// TIA Portal project "Respirator2020_V16" (V16) (continued)
REGION Network 6: Volume/Minute Alarms / Minute Volume Alarms
   RUNG wire#powerrail
      "DirectAnalog_DB_VolumeMinute"(Pulse := "Clock_1Hz", ACK := "Operation".GeneralAck, Reset := "Operation".GeneralReset, Interlock := "Operation".InterlockVolMinute, Delay := T#1000ms, Factor := "OperatingParameters".VolumeMinFactor, AnalogInput := "DataValues".VolumeMinuteValue, SetpointPreAlarmHI := "ProcessData".VolumeMinSetpointPreAlarmHI, SetpointAlarmHI := "ProcessData".VolumeMinSetpointAlarmHI, SetpointPreAlarmLOW := "ProcessData".VolumeMinSetpointPreAlarmLOW, SetpointAlarmLOW := "ProcessData".VolumeMinSetpointAlarmLOW, HysteresisHI := "ProcessData".VolumeMinHysteresisHI, HysteresisLOW := "ProcessData".VolumeMinHysteresisLOW, DisplayPreAlarmHI => "AlarmsRaw".VolumeMinuteDisplayPreAlarmHI, InterlockPreAlarmHI => "AlarmsRaw".VolumeMinuteInterlockPreAlarmHI, DisplayAlarmHI => "AlarmsRaw".VolumeMinuteDisplayAlarmHI, InterlockAlarmHI => "AlarmsRaw".VolumeMinuteInterlockAlarmHI, DisplayPreAlarmLOW => "AlarmsRaw".VolumeMinuteDisplayPreAlarmLOW, InterlockPreAlarmLOW => "AlarmsRaw".VolumeMinuteInterlockPreAlarmLOW, DisplayAlarmLOW => "AlarmsRaw".VolumeMinuteDisplayAlarmLOW, InterlockAlarmLOW => "AlarmsRaw".VolumeMinuteInterlockAlarmLOW, CovertedOutput =>, CalcHysterisHI =>, CalcHysteresisLOW =>, DATOS =>)
   END_RUNG
   // the same network as SCL:
   "DirectAnalog_DB_VolumeMinute"(Pulse := "Clock_1Hz",   // "DirectAnalog"
                           ACK := "Operation".GeneralAck,
                           Reset := "Operation".GeneralReset,
                           Interlock := "Operation".InterlockVolMinute,
                           Delay := T#1000ms,
                           Factor := "OperatingParameters".VolumeMinFactor,
                           AnalogInput := "DataValues".VolumeMinuteValue,
                           SetpointPreAlarmHI := "ProcessData".VolumeMinSetpointPreAlarmHI,
                           SetpointAlarmHI := "ProcessData".VolumeMinSetpointAlarmHI,
                           SetpointPreAlarmLOW := "ProcessData".VolumeMinSetpointPreAlarmLOW,
                           SetpointAlarmLOW := "ProcessData".VolumeMinSetpointAlarmLOW,
                           HysteresisHI := "ProcessData".VolumeMinHysteresisHI,
                           HysteresisLOW := "ProcessData".VolumeMinHysteresisLOW,
                           DisplayPreAlarmHI => "AlarmsRaw".VolumeMinuteDisplayPreAlarmHI,
                           InterlockPreAlarmHI => "AlarmsRaw".VolumeMinuteInterlockPreAlarmHI,
                           DisplayAlarmHI => "AlarmsRaw".VolumeMinuteDisplayAlarmHI,
                           InterlockAlarmHI => "AlarmsRaw".VolumeMinuteInterlockAlarmHI,
                           DisplayPreAlarmLOW => "AlarmsRaw".VolumeMinuteDisplayPreAlarmLOW,
                           InterlockPreAlarmLOW => "AlarmsRaw".VolumeMinuteInterlockPreAlarmLOW,
                           DisplayAlarmLOW => "AlarmsRaw".VolumeMinuteDisplayAlarmLOW,
                           InterlockAlarmLOW => "AlarmsRaw".VolumeMinuteInterlockAlarmLOW);
END_REGION

REGION Network 7: Trigger Alarms
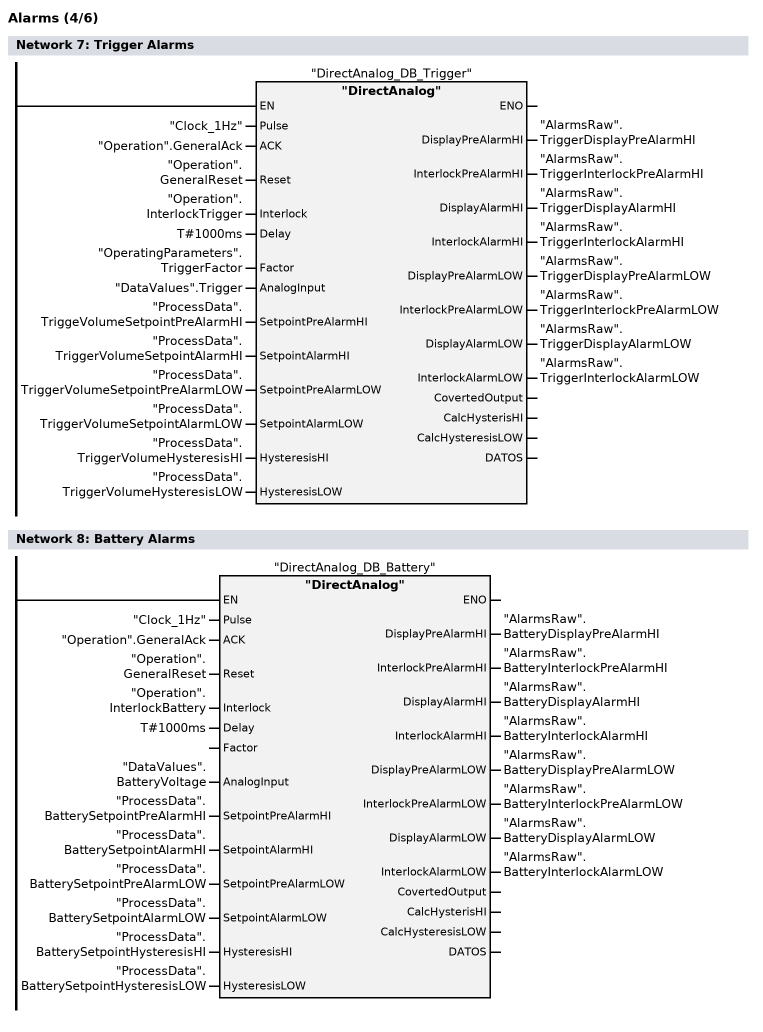
   RUNG wire#powerrail
      "DirectAnalog_DB_Trigger"(Pulse := "Clock_1Hz", ACK := "Operation".GeneralAck, Reset := "Operation".GeneralReset, Interlock := "Operation".InterlockTrigger, Delay := T#1000ms, Factor := "OperatingParameters".TriggerFactor, AnalogInput := "DataValues".Trigger, SetpointPreAlarmHI := "ProcessData".TriggeVolumeSetpointPreAlarmHI, SetpointAlarmHI := "ProcessData".TriggerVolumeSetpointAlarmHI, SetpointPreAlarmLOW := "ProcessData".TriggerVolumeSetpointPreAlarmLOW, SetpointAlarmLOW := "ProcessData".TriggerVolumeSetpointAlarmLOW, HysteresisHI := "ProcessData".TriggerVolumeHysteresisHI, HysteresisLOW := "ProcessData".TriggerVolumeHysteresisLOW, DisplayPreAlarmHI => "AlarmsRaw".TriggerDisplayPreAlarmHI, InterlockPreAlarmHI => "AlarmsRaw".TriggerInterlockPreAlarmHI, DisplayAlarmHI => "AlarmsRaw".TriggerDisplayAlarmHI, InterlockAlarmHI => "AlarmsRaw".TriggerInterlockAlarmHI, DisplayPreAlarmLOW => "AlarmsRaw".TriggerDisplayPreAlarmLOW, InterlockPreAlarmLOW => "AlarmsRaw".TriggerInterlockPreAlarmLOW, DisplayAlarmLOW => "AlarmsRaw".TriggerDisplayAlarmLOW, InterlockAlarmLOW => "AlarmsRaw".TriggerInterlockAlarmLOW, CovertedOutput =>, CalcHysterisHI =>, CalcHysteresisLOW =>, DATOS =>)
   END_RUNG
   // the same network as SCL:
   "DirectAnalog_DB_Trigger"(Pulse := "Clock_1Hz",   // "DirectAnalog"
                           ACK := "Operation".GeneralAck,
                           Reset := "Operation".GeneralReset,
                           Interlock := "Operation".InterlockTrigger,
                           Delay := T#1000ms,
                           Factor := "OperatingParameters".TriggerFactor,
                           AnalogInput := "DataValues".Trigger,
                           SetpointPreAlarmHI := "ProcessData".TriggeVolumeSetpointPreAlarmHI,
                           SetpointAlarmHI := "ProcessData".TriggerVolumeSetpointAlarmHI,
                           SetpointPreAlarmLOW := "ProcessData".TriggerVolumeSetpointPreAlarmLOW,
                           SetpointAlarmLOW := "ProcessData".TriggerVolumeSetpointAlarmLOW,
                           HysteresisHI := "ProcessData".TriggerVolumeHysteresisHI,
                           HysteresisLOW := "ProcessData".TriggerVolumeHysteresisLOW,
                           DisplayPreAlarmHI => "AlarmsRaw".TriggerDisplayPreAlarmHI,
                           InterlockPreAlarmHI => "AlarmsRaw".TriggerInterlockPreAlarmHI,
                           DisplayAlarmHI => "AlarmsRaw".TriggerDisplayAlarmHI,
                           InterlockAlarmHI => "AlarmsRaw".TriggerInterlockAlarmHI,
                           DisplayPreAlarmLOW => "AlarmsRaw".TriggerDisplayPreAlarmLOW,
                           InterlockPreAlarmLOW => "AlarmsRaw".TriggerInterlockPreAlarmLOW,
                           DisplayAlarmLOW => "AlarmsRaw".TriggerDisplayAlarmLOW,
                           InterlockAlarmLOW => "AlarmsRaw".TriggerInterlockAlarmLOW);
END_REGION

REGION Network 8: Battery Alarms
   RUNG wire#powerrail
      "DirectAnalog_DB_Battery"(Pulse := "Clock_1Hz", ACK := "Operation".GeneralAck, Reset := "Operation".GeneralReset, Interlock := "Operation".InterlockBattery, Delay := T#1000ms, Factor :=, AnalogInput := "DataValues".BatteryVoltage, SetpointPreAlarmHI := "ProcessData".BatterySetpointPreAlarmHI, SetpointAlarmHI := "ProcessData".BatterySetpointAlarmHI, SetpointPreAlarmLOW := "ProcessData".BatterySetpointPreAlarmLOW, SetpointAlarmLOW := "ProcessData".BatterySetpointAlarmLOW, HysteresisHI := "ProcessData".BatterySetpointHysteresisHI, HysteresisLOW := "ProcessData".BatterySetpointHysteresisLOW, DisplayPreAlarmHI => "AlarmsRaw".BatteryDisplayPreAlarmHI, InterlockPreAlarmHI => "AlarmsRaw".BatteryInterlockPreAlarmHI, DisplayAlarmHI => "AlarmsRaw".BatteryDisplayAlarmHI, InterlockAlarmHI => "AlarmsRaw".BatteryInterlockAlarmHI, DisplayPreAlarmLOW => "AlarmsRaw".BatteryDisplayPreAlarmLOW, InterlockPreAlarmLOW => "AlarmsRaw".BatteryInterlockPreAlarmLOW, DisplayAlarmLOW => "AlarmsRaw".BatteryDisplayAlarmLOW, InterlockAlarmLOW => "AlarmsRaw".BatteryInterlockAlarmLOW, CovertedOutput =>, CalcHysterisHI =>, CalcHysteresisLOW =>, DATOS =>)
   END_RUNG
   // the same network as SCL:
   "DirectAnalog_DB_Battery"(Pulse := "Clock_1Hz",   // "DirectAnalog"
                           ACK := "Operation".GeneralAck,
                           Reset := "Operation".GeneralReset,
                           Interlock := "Operation".InterlockBattery,
                           Delay := T#1000ms,
                           AnalogInput := "DataValues".BatteryVoltage,
                           SetpointPreAlarmHI := "ProcessData".BatterySetpointPreAlarmHI,
                           SetpointAlarmHI := "ProcessData".BatterySetpointAlarmHI,
                           SetpointPreAlarmLOW := "ProcessData".BatterySetpointPreAlarmLOW,
                           SetpointAlarmLOW := "ProcessData".BatterySetpointAlarmLOW,
                           HysteresisHI := "ProcessData".BatterySetpointHysteresisHI,
                           HysteresisLOW := "ProcessData".BatterySetpointHysteresisLOW,
                           DisplayPreAlarmHI => "AlarmsRaw".BatteryDisplayPreAlarmHI,
                           InterlockPreAlarmHI => "AlarmsRaw".BatteryInterlockPreAlarmHI,
                           DisplayAlarmHI => "AlarmsRaw".BatteryDisplayAlarmHI,
                           InterlockAlarmHI => "AlarmsRaw".BatteryInterlockAlarmHI,
                           DisplayPreAlarmLOW => "AlarmsRaw".BatteryDisplayPreAlarmLOW,
                           InterlockPreAlarmLOW => "AlarmsRaw".BatteryInterlockPreAlarmLOW,
                           DisplayAlarmLOW => "AlarmsRaw".BatteryDisplayAlarmLOW,
                           InterlockAlarmLOW => "AlarmsRaw".BatteryInterlockAlarmLOW);
END_REGION

REGION Network 9: ALARM-0 Packing
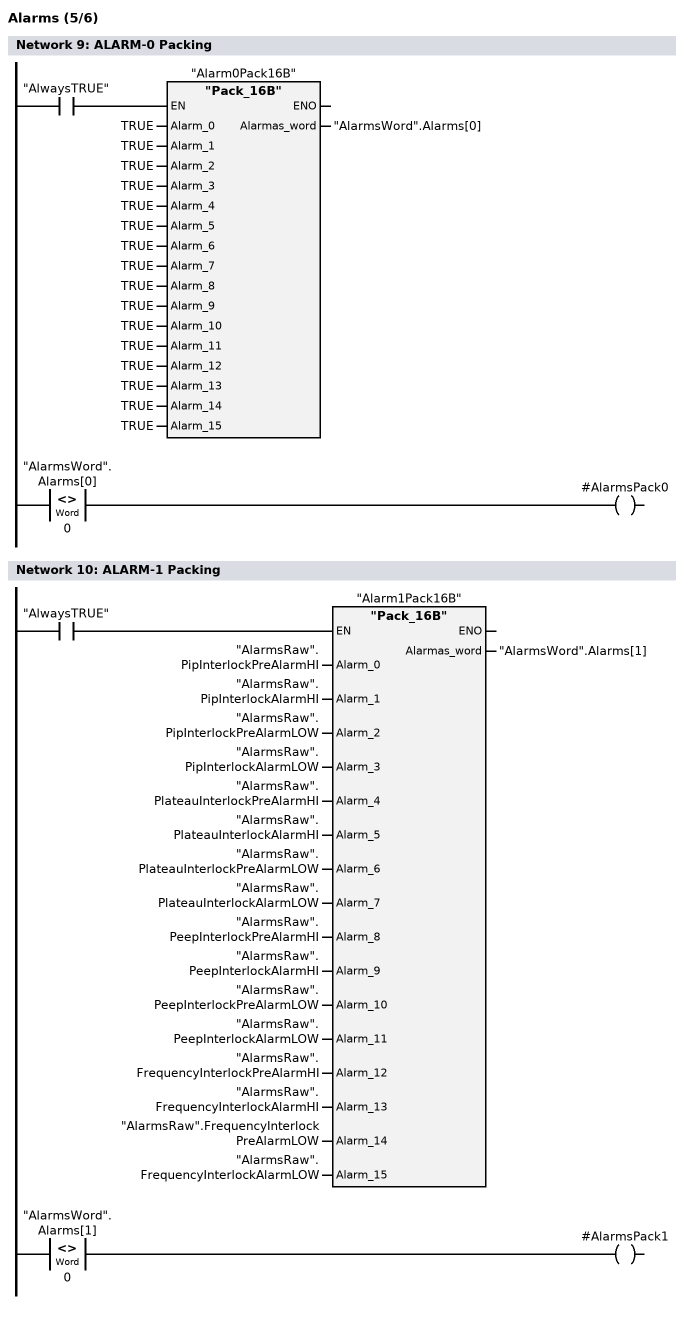
   RUNG wire#powerrail
      Contact( "AlwaysTRUE" )
      "Alarm0Pack16B"(Alarm_0 := TRUE, Alarm_1 := TRUE, Alarm_2 := TRUE, Alarm_3 := TRUE, Alarm_4 := TRUE, Alarm_5 := TRUE, Alarm_6 := TRUE, Alarm_7 := TRUE, Alarm_8 := TRUE, Alarm_9 := TRUE, Alarm_10 := TRUE, Alarm_11 := TRUE, Alarm_12 := TRUE, Alarm_13 := TRUE, Alarm_14 := TRUE, Alarm_15 := TRUE, Alarmas_word => "AlarmsWord".Alarms[0])
   END_RUNG
   RUNG wire#powerrail
      { S7_Templates := "SrcType := Word" } NE_Contact(in1 := "AlarmsWord".Alarms[0], in2 := 0)
      Coil( #AlarmsPack0 )
   END_RUNG
   // the same network as SCL:
   IF "AlwaysTRUE" THEN
       "Alarm0Pack16B"(Alarm_0 := TRUE,   // "Pack_16B"
                       Alarm_1 := TRUE,
                       Alarm_2 := TRUE,
                       Alarm_3 := TRUE,
                       Alarm_4 := TRUE,
                       Alarm_5 := TRUE,
                       Alarm_6 := TRUE,
                       Alarm_7 := TRUE,
                       Alarm_8 := TRUE,
                       Alarm_9 := TRUE,
                       Alarm_10 := TRUE,
                       Alarm_11 := TRUE,
                       Alarm_12 := TRUE,
                       Alarm_13 := TRUE,
                       Alarm_14 := TRUE,
                       Alarm_15 := TRUE,
                       Alarmas_word => "AlarmsWord".Alarms[0]);
   END_IF;
   #AlarmsPack0 := "AlarmsWord".Alarms[0] <> 0;
END_REGION

REGION Network 10: ALARM-1 Packing
   RUNG wire#powerrail
      Contact( "AlwaysTRUE" )
      "Alarm1Pack16B"(Alarm_0 := "AlarmsRaw".PipInterlockPreAlarmHI, Alarm_1 := "AlarmsRaw".PipInterlockAlarmHI, Alarm_2 := "AlarmsRaw".PipInterlockPreAlarmLOW, Alarm_3 := "AlarmsRaw".PipInterlockAlarmLOW, Alarm_4 := "AlarmsRaw".PlateauInterlockPreAlarmHI, Alarm_5 := "AlarmsRaw".PlateauInterlockAlarmHI, Alarm_6 := "AlarmsRaw".PlateauInterlockPreAlarmLOW, Alarm_7 := "AlarmsRaw".PlateauInterlockAlarmLOW, Alarm_8 := "AlarmsRaw".PeepInterlockPreAlarmHI, Alarm_9 := "AlarmsRaw".PeepInterlockAlarmHI, Alarm_10 := "AlarmsRaw".PeepInterlockPreAlarmLOW, Alarm_11 := "AlarmsRaw".PeepInterlockAlarmLOW, Alarm_12 := "AlarmsRaw".FrequencyInterlockPreAlarmHI, Alarm_13 := "AlarmsRaw".FrequencyInterlockAlarmHI, Alarm_14 := "AlarmsRaw".FrequencyInterlockPreAlarmLOW, Alarm_15 := "AlarmsRaw".FrequencyInterlockAlarmLOW, Alarmas_word => "AlarmsWord".Alarms[1])
   END_RUNG
   RUNG wire#powerrail
      { S7_Templates := "SrcType := Word" } NE_Contact(in1 := "AlarmsWord".Alarms[1], in2 := 0)
      Coil( #AlarmsPack1 )
   END_RUNG
   // the same network as SCL:
   IF "AlwaysTRUE" THEN
       "Alarm1Pack16B"(Alarm_0 := "AlarmsRaw".PipInterlockPreAlarmHI,   // "Pack_16B"
                       Alarm_1 := "AlarmsRaw".PipInterlockAlarmHI,
                       Alarm_2 := "AlarmsRaw".PipInterlockPreAlarmLOW,
                       Alarm_3 := "AlarmsRaw".PipInterlockAlarmLOW,
                       Alarm_4 := "AlarmsRaw".PlateauInterlockPreAlarmHI,
                       Alarm_5 := "AlarmsRaw".PlateauInterlockAlarmHI,
                       Alarm_6 := "AlarmsRaw".PlateauInterlockPreAlarmLOW,
                       Alarm_7 := "AlarmsRaw".PlateauInterlockAlarmLOW,
                       Alarm_8 := "AlarmsRaw".PeepInterlockPreAlarmHI,
                       Alarm_9 := "AlarmsRaw".PeepInterlockAlarmHI,
                       Alarm_10 := "AlarmsRaw".PeepInterlockPreAlarmLOW,
                       Alarm_11 := "AlarmsRaw".PeepInterlockAlarmLOW,
                       Alarm_12 := "AlarmsRaw".FrequencyInterlockPreAlarmHI,
                       Alarm_13 := "AlarmsRaw".FrequencyInterlockAlarmHI,
                       Alarm_14 := "AlarmsRaw".FrequencyInterlockPreAlarmLOW,
                       Alarm_15 := "AlarmsRaw".FrequencyInterlockAlarmLOW,
                       Alarmas_word => "AlarmsWord".Alarms[1]);
   END_IF;
   #AlarmsPack1 := "AlarmsWord".Alarms[1] <> 0;
END_REGION

REGION Network 11: ALARM-2 Packing
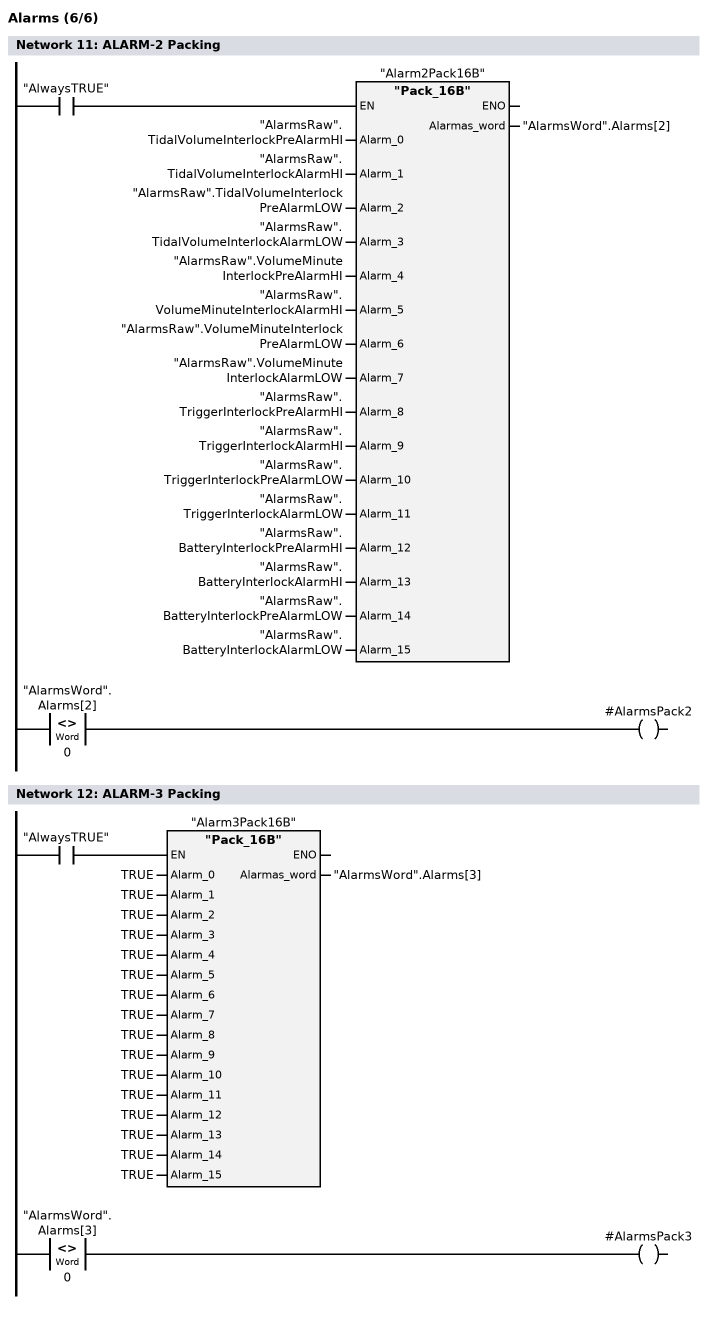
   RUNG wire#powerrail
      Contact( "AlwaysTRUE" )
      "Alarm2Pack16B"(Alarm_0 := "AlarmsRaw".TidalVolumeInterlockPreAlarmHI, Alarm_1 := "AlarmsRaw".TidalVolumeInterlockAlarmHI, Alarm_2 := "AlarmsRaw".TidalVolumeInterlockPreAlarmLOW, Alarm_3 := "AlarmsRaw".TidalVolumeInterlockAlarmLOW, Alarm_4 := "AlarmsRaw".VolumeMinuteInterlockPreAlarmHI, Alarm_5 := "AlarmsRaw".VolumeMinuteInterlockAlarmHI, Alarm_6 := "AlarmsRaw".VolumeMinuteInterlockPreAlarmLOW, Alarm_7 := "AlarmsRaw".VolumeMinuteInterlockAlarmLOW, Alarm_8 := "AlarmsRaw".TriggerInterlockPreAlarmHI, Alarm_9 := "AlarmsRaw".TriggerInterlockAlarmHI, Alarm_10 := "AlarmsRaw".TriggerInterlockPreAlarmLOW, Alarm_11 := "AlarmsRaw".TriggerInterlockAlarmLOW, Alarm_12 := "AlarmsRaw".BatteryInterlockPreAlarmHI, Alarm_13 := "AlarmsRaw".BatteryInterlockAlarmHI, Alarm_14 := "AlarmsRaw".BatteryInterlockPreAlarmLOW, Alarm_15 := "AlarmsRaw".BatteryInterlockAlarmLOW, Alarmas_word => "AlarmsWord".Alarms[2])
   END_RUNG
   RUNG wire#powerrail
      { S7_Templates := "SrcType := Word" } NE_Contact(in1 := "AlarmsWord".Alarms[2], in2 := 0)
      Coil( #AlarmsPack2 )
   END_RUNG
   // the same network as SCL:
   IF "AlwaysTRUE" THEN
       "Alarm2Pack16B"(Alarm_0 := "AlarmsRaw".TidalVolumeInterlockPreAlarmHI,   // "Pack_16B"
                       Alarm_1 := "AlarmsRaw".TidalVolumeInterlockAlarmHI,
                       Alarm_2 := "AlarmsRaw".TidalVolumeInterlockPreAlarmLOW,
                       Alarm_3 := "AlarmsRaw".TidalVolumeInterlockAlarmLOW,
                       Alarm_4 := "AlarmsRaw".VolumeMinuteInterlockPreAlarmHI,
                       Alarm_5 := "AlarmsRaw".VolumeMinuteInterlockAlarmHI,
                       Alarm_6 := "AlarmsRaw".VolumeMinuteInterlockPreAlarmLOW,
                       Alarm_7 := "AlarmsRaw".VolumeMinuteInterlockAlarmLOW,
                       Alarm_8 := "AlarmsRaw".TriggerInterlockPreAlarmHI,
                       Alarm_9 := "AlarmsRaw".TriggerInterlockAlarmHI,
                       Alarm_10 := "AlarmsRaw".TriggerInterlockPreAlarmLOW,
                       Alarm_11 := "AlarmsRaw".TriggerInterlockAlarmLOW,
                       Alarm_12 := "AlarmsRaw".BatteryInterlockPreAlarmHI,
                       Alarm_13 := "AlarmsRaw".BatteryInterlockAlarmHI,
                       Alarm_14 := "AlarmsRaw".BatteryInterlockPreAlarmLOW,
                       Alarm_15 := "AlarmsRaw".BatteryInterlockAlarmLOW,
                       Alarmas_word => "AlarmsWord".Alarms[2]);
   END_IF;
   #AlarmsPack2 := "AlarmsWord".Alarms[2] <> 0;
END_REGION

REGION Network 12: ALARM-3 Packing
   RUNG wire#powerrail
      Contact( "AlwaysTRUE" )
      "Alarm3Pack16B"(Alarm_0 := TRUE, Alarm_1 := TRUE, Alarm_2 := TRUE, Alarm_3 := TRUE, Alarm_4 := TRUE, Alarm_5 := TRUE, Alarm_6 := TRUE, Alarm_7 := TRUE, Alarm_8 := TRUE, Alarm_9 := TRUE, Alarm_10 := TRUE, Alarm_11 := TRUE, Alarm_12 := TRUE, Alarm_13 := TRUE, Alarm_14 := TRUE, Alarm_15 := TRUE, Alarmas_word => "AlarmsWord".Alarms[3])
   END_RUNG
   RUNG wire#powerrail
      { S7_Templates := "SrcType := Word" } NE_Contact(in1 := "AlarmsWord".Alarms[3], in2 := 0)
      Coil( #AlarmsPack3 )
   END_RUNG
   // the same network as SCL:
   IF "AlwaysTRUE" THEN
       "Alarm3Pack16B"(Alarm_0 := TRUE,   // "Pack_16B"
                       Alarm_1 := TRUE,
                       Alarm_2 := TRUE,
                       Alarm_3 := TRUE,
                       Alarm_4 := TRUE,
                       Alarm_5 := TRUE,
                       Alarm_6 := TRUE,
                       Alarm_7 := TRUE,
                       Alarm_8 := TRUE,
                       Alarm_9 := TRUE,
                       Alarm_10 := TRUE,
                       Alarm_11 := TRUE,
                       Alarm_12 := TRUE,
                       Alarm_13 := TRUE,
                       Alarm_14 := TRUE,
                       Alarm_15 := TRUE,
                       Alarmas_word => "AlarmsWord".Alarms[3]);
   END_IF;
   #AlarmsPack3 := "AlarmsWord".Alarms[3] <> 0;
END_REGION
END_FUNCTION_BLOCK

// folder: 4_ProcessControl

FUNCTION_BLOCK "0_ProcessControl"   // FB40, LAD
TITLE = Proccess Control
{ S7_Optimized_Access := 'TRUE' }
AUTHOR : JL_Cristobal_2020
VERSION : 0.1
   VAR
      REFrecuencyPlus : Bool;
      REFrecuencyMinus : Bool;
      REPeakPlus : Bool;
      REPeakMinus : Bool;
      REPeepPlus : Bool;
      REPeepMinus : Bool;
      REPowerError : Bool;
      test : Bool;
   END_VAR
BEGIN

REGION Network 1: Motor Enable
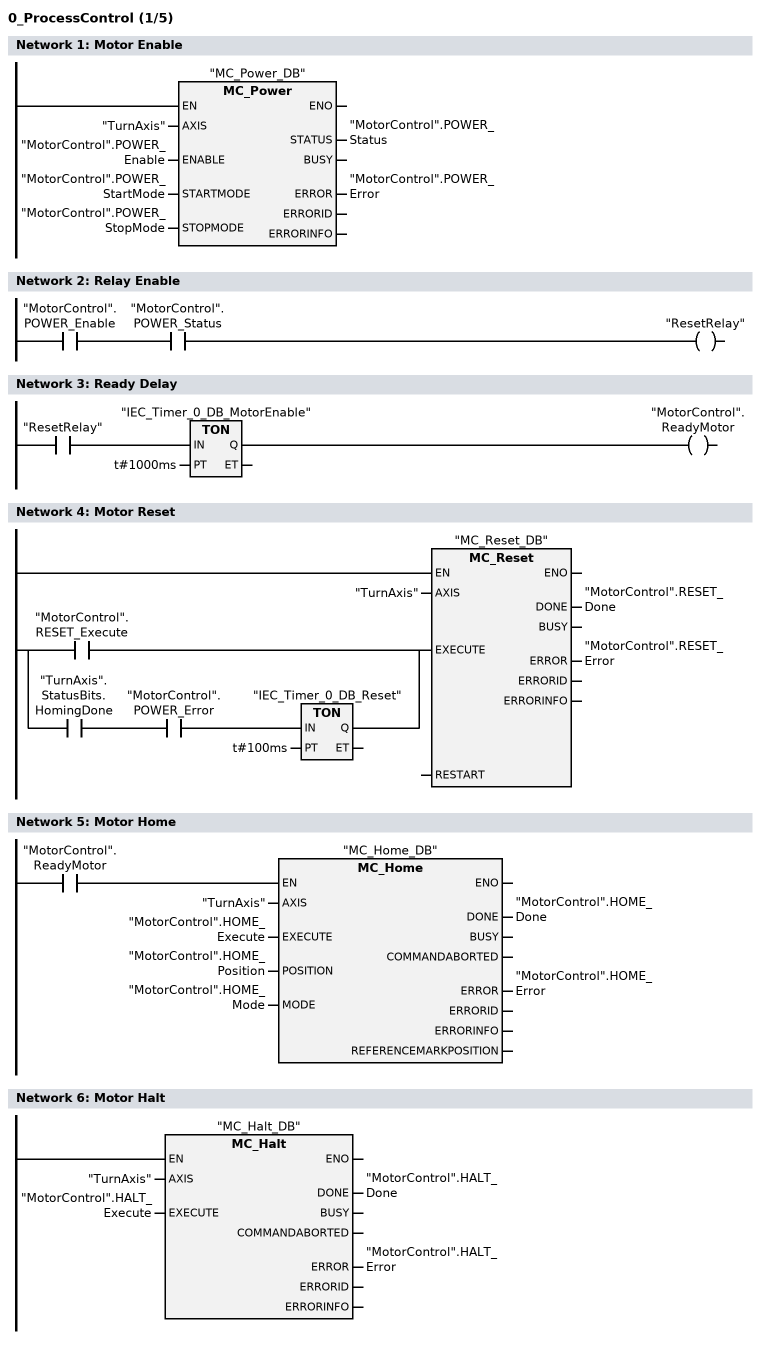
   "MC_Power_DB"(Axis := "TurnAxis",   // MC_Power
                 Enable := "MotorControl".POWER_Enable,
                 StartMode := "MotorControl".POWER_StartMode,
                 StopMode := "MotorControl".POWER_StopMode,
                 Status => "MotorControl".POWER_Status,
                 Error => "MotorControl".POWER_Error);
END_REGION

REGION Network 2: Relay Enable
   RUNG wire#powerrail
      Contact( "MotorControl".POWER_Enable )
      Contact( "MotorControl".POWER_Status )
      Coil( "ResetRelay" )
   END_RUNG
   // the same network as SCL:
   "ResetRelay" := "MotorControl".POWER_Enable AND "MotorControl".POWER_Status;
END_REGION

REGION Network 3: Ready Delay
   "IEC_Timer_0_DB_MotorEnable".TON(IN := "ResetRelay", PT := t#1000ms);
   "MotorControl".ReadyMotor := "IEC_Timer_0_DB_MotorEnable".Q;
END_REGION

REGION Network 4: Motor Reset
   "IEC_Timer_0_DB_Reset".TON(IN := "TurnAxis".StatusBits.HomingDone AND "MotorControl".POWER_Error,
                           PT := t#100ms);
   "MC_Reset_DB"(Axis := "TurnAxis",   // MC_Reset
                 Execute := "MotorControl".RESET_Execute OR "IEC_Timer_0_DB_Reset".Q,
                 Done => "MotorControl".RESET_Done,
                 Error => "MotorControl".RESET_Error);
END_REGION

REGION Network 5: Motor Home
   IF "MotorControl".ReadyMotor THEN
       "MC_Home_DB"(Axis := "TurnAxis",   // MC_Home
                    Execute := "MotorControl".HOME_Execute,
                    Position := "MotorControl".HOME_Position,
                    Mode := "MotorControl".HOME_Mode,
                    Done => "MotorControl".HOME_Done,
                    Error => "MotorControl".HOME_Error);
   END_IF;
END_REGION

REGION Network 6: Motor Halt
   "MC_Halt_DB"(Axis := "TurnAxis",   // MC_Halt
                Execute := "MotorControl".HALT_Execute,
                Done => "MotorControl".HALT_Done,
                Error => "MotorControl".HALT_Error);
END_REGION

REGION Network 7: Motor Move Absolute
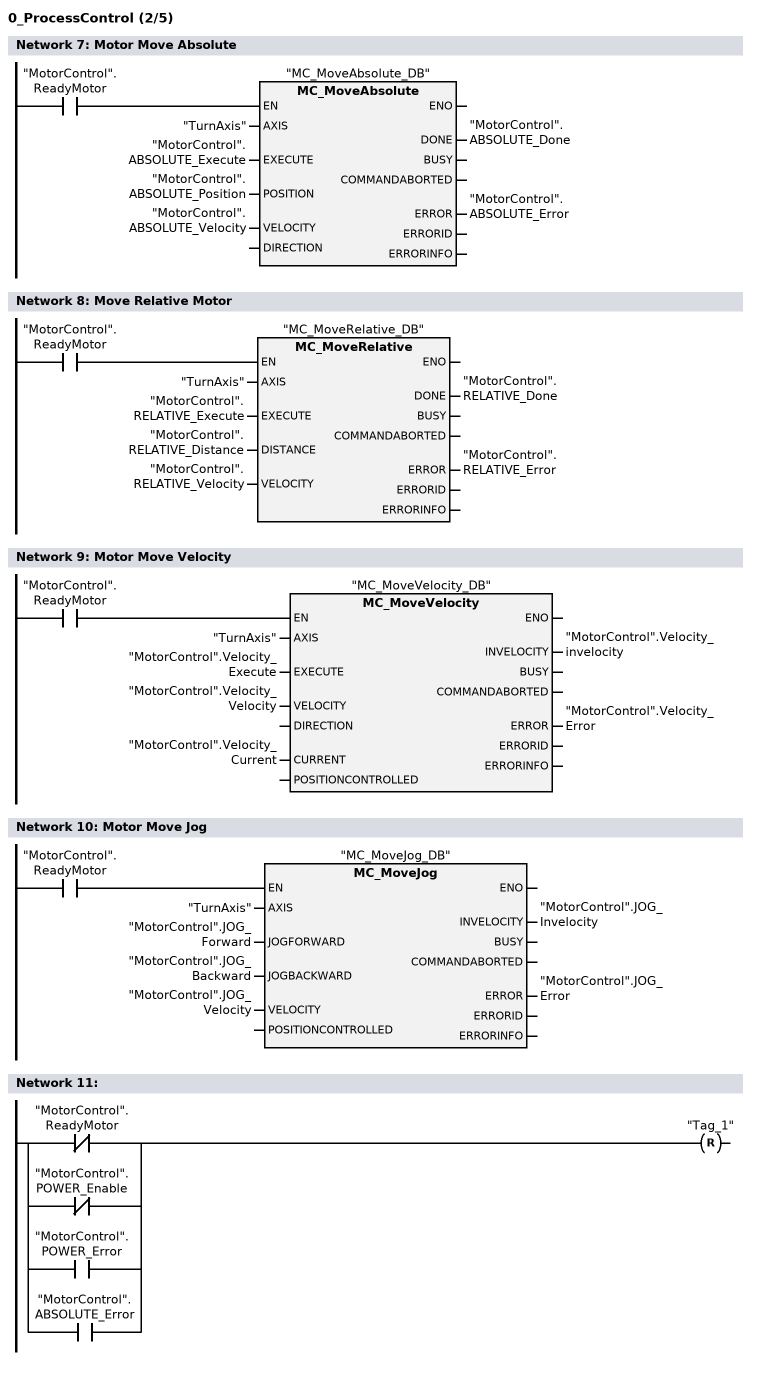
   IF "MotorControl".ReadyMotor THEN
       "MC_MoveAbsolute_DB"(Axis := "TurnAxis",   // MC_MoveAbsolute
                            Execute := "MotorControl".ABSOLUTE_Execute,
                            Position := "MotorControl".ABSOLUTE_Position,
                            Velocity := "MotorControl".ABSOLUTE_Velocity,
                            Done => "MotorControl".ABSOLUTE_Done,
                            Error => "MotorControl".ABSOLUTE_Error);
   END_IF;
END_REGION

REGION Network 8: Move Relative Motor
   IF "MotorControl".ReadyMotor THEN
       "MC_MoveRelative_DB"(Axis := "TurnAxis",   // MC_MoveRelative
                            Execute := "MotorControl".RELATIVE_Execute,
                            Distance := "MotorControl".RELATIVE_Distance,
                            Velocity := "MotorControl".RELATIVE_Velocity,
                            Done => "MotorControl".RELATIVE_Done,
                            Error => "MotorControl".RELATIVE_Error);
   END_IF;
END_REGION

REGION Network 9: Motor Move Velocity
   IF "MotorControl".ReadyMotor THEN
       "MC_MoveVelocity_DB"(Axis := "TurnAxis",   // MC_MoveVelocity
                            Execute := "MotorControl".Velocity_Execute,
                            Velocity := "MotorControl".Velocity_Velocity,
                            Current := "MotorControl".Velocity_Current,
                            InVelocity => "MotorControl".Velocity_invelocity,
                            Error => "MotorControl".Velocity_Error);
   END_IF;
END_REGION

REGION Network 10: Motor Move Jog
   IF "MotorControl".ReadyMotor THEN
       "MC_MoveJog_DB"(Axis := "TurnAxis",   // MC_MoveJog
                       JogForward := "MotorControl".JOG_Forward,
                       JogBackward := "MotorControl".JOG_Backward,
                       Velocity := "MotorControl".JOG_Velocity,
                       InVelocity => "MotorControl".JOG_Invelocity,
                       Error => "MotorControl".JOG_Error);
   END_IF;
END_REGION

REGION Network 11
   RUNG wire#powerrail
      I_Contact( "MotorControl".ReadyMotor )
      wire#w1
      R_Coil( "Tag_1" )
   END_RUNG
   RUNG wire#powerrail
      I_Contact( "MotorControl".POWER_Enable )
   END_RUNG wire#w1
   RUNG wire#powerrail
      Contact( "MotorControl".POWER_Error )
   END_RUNG wire#w1
   RUNG wire#powerrail
      Contact( "MotorControl".ABSOLUTE_Error )
   END_RUNG wire#w1
   // the same network as SCL:
   IF NOT "MotorControl".ReadyMotor OR NOT "MotorControl".POWER_Enable OR "MotorControl".POWER_Error OR "MotorControl".ABSOLUTE_Error THEN
       "Tag_1" := FALSE;
   END_IF;
END_REGION

REGION Network 12: test
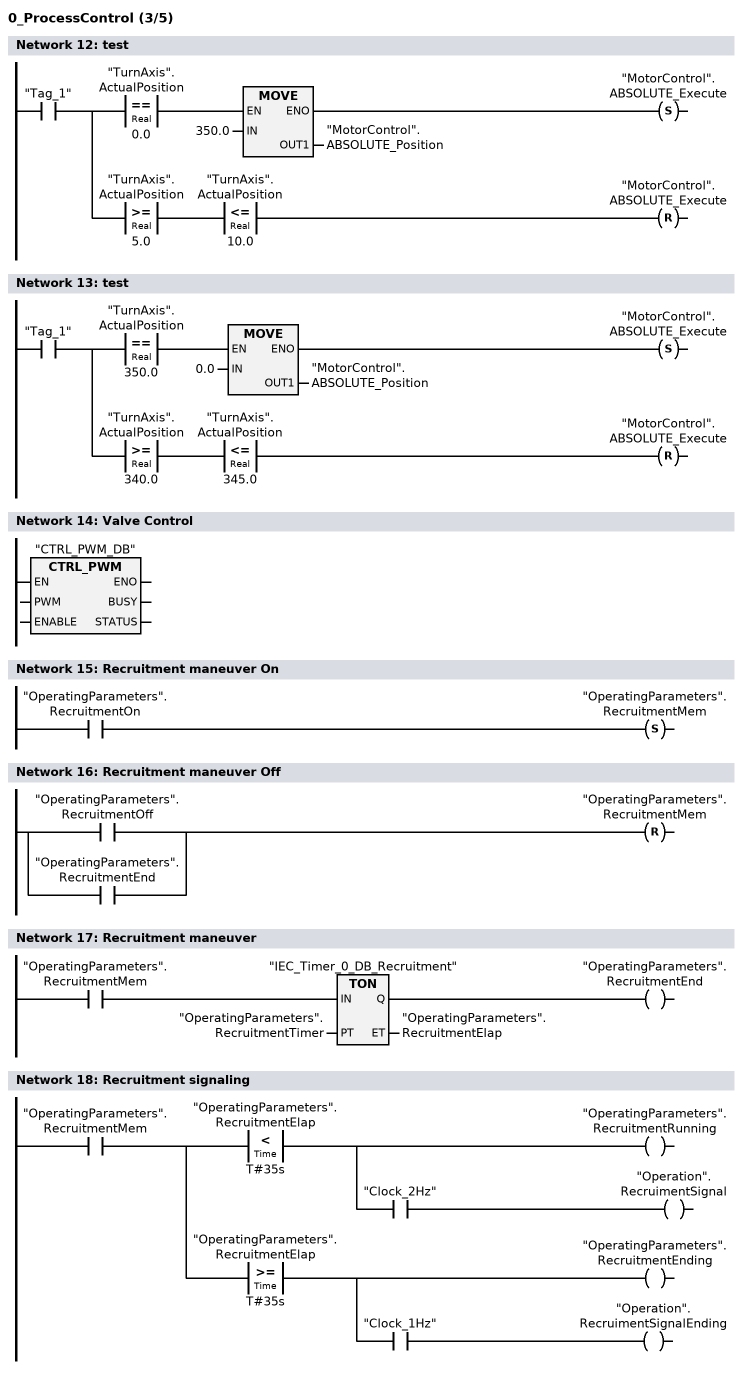
   RUNG wire#powerrail
      Contact( "Tag_1" )
      wire#w1
      { S7_Templates := "SrcType := Real" } EQ_Contact(in1 := "TurnAxis".ActualPosition, in2 := 0.0)
      Move(in := 350.0, out1 => "MotorControl".ABSOLUTE_Position)
      S_Coil( "MotorControl".ABSOLUTE_Execute )
   END_RUNG
   RUNG wire#w1
      { S7_Templates := "SrcType := Real" } GE_Contact(in1 := "TurnAxis".ActualPosition, in2 := 5.0)
      { S7_Templates := "SrcType := Real" } LE_Contact(in1 := "TurnAxis".ActualPosition, in2 := 10.0)
      R_Coil( "MotorControl".ABSOLUTE_Execute )
   END_RUNG
   // the same network as SCL:
   IF "Tag_1" AND ("TurnAxis".ActualPosition = 0.0) THEN
       "MotorControl".ABSOLUTE_Position := 350.0;
       "MotorControl".ABSOLUTE_Execute := TRUE;
   END_IF;
   IF "Tag_1" AND ("TurnAxis".ActualPosition >= 5.0) AND ("TurnAxis".ActualPosition <= 10.0) THEN
       "MotorControl".ABSOLUTE_Execute := FALSE;
   END_IF;
END_REGION

REGION Network 13: test
   RUNG wire#powerrail
      Contact( "Tag_1" )
      wire#w1
      { S7_Templates := "SrcType := Real" } EQ_Contact(in1 := "TurnAxis".ActualPosition, in2 := 350.0)
      Move(in := 0.0, out1 => "MotorControl".ABSOLUTE_Position)
      S_Coil( "MotorControl".ABSOLUTE_Execute )
   END_RUNG
   RUNG wire#w1
      { S7_Templates := "SrcType := Real" } GE_Contact(in1 := "TurnAxis".ActualPosition, in2 := 340.0)
      { S7_Templates := "SrcType := Real" } LE_Contact(in1 := "TurnAxis".ActualPosition, in2 := 345.0)
      R_Coil( "MotorControl".ABSOLUTE_Execute )
   END_RUNG
   // the same network as SCL:
   IF "Tag_1" AND ("TurnAxis".ActualPosition = 350.0) THEN
       "MotorControl".ABSOLUTE_Position := 0.0;
       "MotorControl".ABSOLUTE_Execute := TRUE;
   END_IF;
   IF "Tag_1" AND ("TurnAxis".ActualPosition >= 340.0) AND ("TurnAxis".ActualPosition <= 345.0) THEN
       "MotorControl".ABSOLUTE_Execute := FALSE;
   END_IF;
END_REGION

REGION Network 14: Valve Control
   "CTRL_PWM_DB"();   // CTRL_PWM
END_REGION

REGION Network 15: Recruitment maneuver On
   RUNG wire#powerrail
      Contact( "OperatingParameters".RecruitmentOn )
      S_Coil( "OperatingParameters".RecruitmentMem )
   END_RUNG
   // the same network as SCL:
   IF "OperatingParameters".RecruitmentOn THEN "OperatingParameters".RecruitmentMem := TRUE; END_IF;
END_REGION

REGION Network 16: Recruitment maneuver Off
   RUNG wire#powerrail
      Contact( "OperatingParameters".RecruitmentOff )
      wire#w1
      R_Coil( "OperatingParameters".RecruitmentMem )
   END_RUNG
   RUNG wire#powerrail
      Contact( "OperatingParameters".RecruitmentEnd )
   END_RUNG wire#w1
   // the same network as SCL:
   IF "OperatingParameters".RecruitmentOff OR "OperatingParameters".RecruitmentEnd THEN
       "OperatingParameters".RecruitmentMem := FALSE;
   END_IF;
END_REGION

REGION Network 17: Recruitment maneuver
   "IEC_Timer_0_DB_Recruitment".TON(IN := "OperatingParameters".RecruitmentMem,
                           PT := "OperatingParameters".RecruitmentTimer,
                           ET => "OperatingParameters".RecruitmentElap);
   "OperatingParameters".RecruitmentEnd := "IEC_Timer_0_DB_Recruitment".Q;
END_REGION

REGION Network 18: Recruitment signaling
   RUNG wire#powerrail
      Contact( "OperatingParameters".RecruitmentMem )
      wire#w1
      { S7_Templates := "SrcType := Time" } LT_Contact(in1 := "OperatingParameters".RecruitmentElap, in2 := T#35s)
      wire#w2
      Coil( "OperatingParameters".RecruitmentRunning )
   END_RUNG
   RUNG wire#w2
      Contact( "Clock_2Hz" )
      Coil( "Operation".RecruimentSignal )
   END_RUNG
   RUNG wire#w1
      { S7_Templates := "SrcType := Time" } GE_Contact(in1 := "OperatingParameters".RecruitmentElap, in2 := T#35s)
      wire#w3
      Coil( "OperatingParameters".RecruitmentEnding )
   END_RUNG
   RUNG wire#w3
      Contact( "Clock_1Hz" )
      Coil( "Operation".RecruimentSignalEnding )
   END_RUNG
   // the same network as SCL:
   "OperatingParameters".RecruitmentRunning := "OperatingParameters".RecruitmentMem AND ("OperatingParameters".RecruitmentElap < T#35s);
   "Operation".RecruimentSignal := "OperatingParameters".RecruitmentRunning AND "Clock_2Hz";
   "OperatingParameters".RecruitmentEnding := "OperatingParameters".RecruitmentMem AND ("OperatingParameters".RecruitmentElap >= T#35s);
   "Operation".RecruimentSignalEnding := "OperatingParameters".RecruitmentEnding AND "Clock_1Hz";
END_REGION

REGION Network 19: Multi point PID Switcher
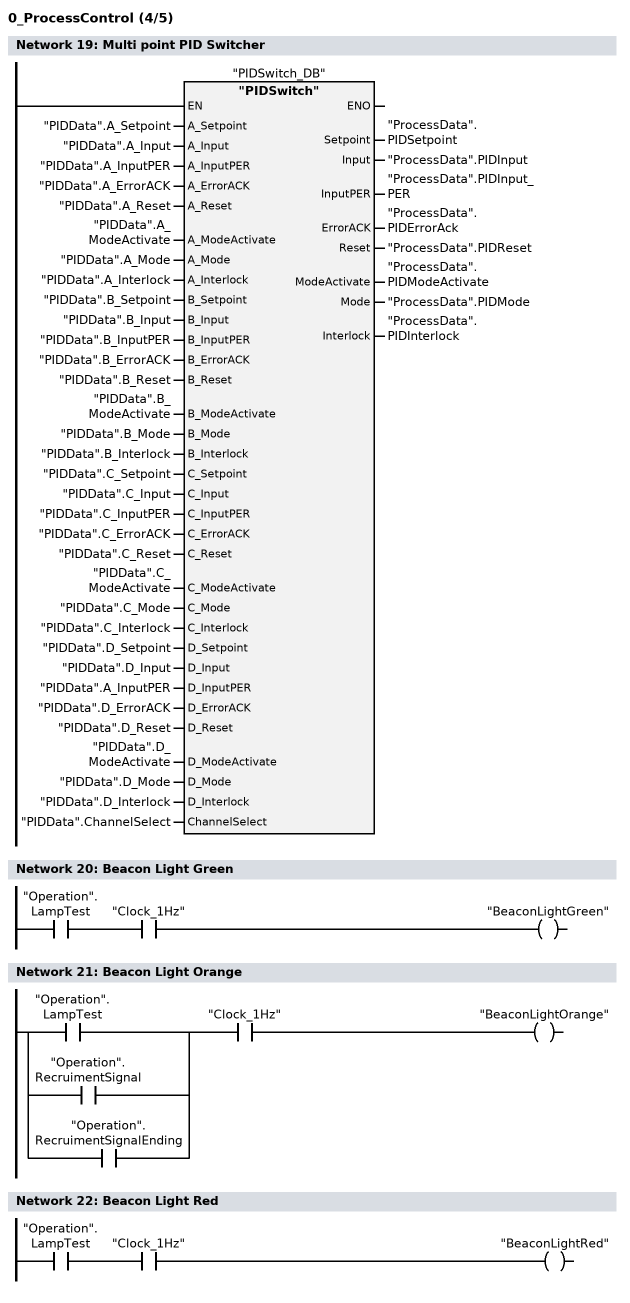
   RUNG wire#powerrail
      "PIDSwitch_DB"(A_Setpoint := "PIDData".A_Setpoint, A_Input := "PIDData".A_Input, A_InputPER := "PIDData".A_InputPER, A_ErrorACK := "PIDData".A_ErrorACK, A_Reset := "PIDData".A_Reset, A_ModeActivate := "PIDData".A_ModeActivate, A_Mode := "PIDData".A_Mode, A_Interlock := "PIDData".A_Interlock, B_Setpoint := "PIDData".B_Setpoint, B_Input := "PIDData".B_Input, B_InputPER := "PIDData".B_InputPER, B_ErrorACK := "PIDData".B_ErrorACK, B_Reset := "PIDData".B_Reset, B_ModeActivate := "PIDData".B_ModeActivate, B_Mode := "PIDData".B_Mode, B_Interlock := "PIDData".B_Interlock, C_Setpoint := "PIDData".C_Setpoint, C_Input := "PIDData".C_Input, C_InputPER := "PIDData".C_InputPER, C_ErrorACK := "PIDData".C_ErrorACK, C_Reset := "PIDData".C_Reset, C_ModeActivate := "PIDData".C_ModeActivate, C_Mode := "PIDData".C_Mode, C_Interlock := "PIDData".C_Interlock, D_Setpoint := "PIDData".D_Setpoint, D_Input := "PIDData".D_Input, D_InputPER := "PIDData".A_InputPER, D_ErrorACK := "PIDData".D_ErrorACK, D_Reset := "PIDData".D_Reset, D_ModeActivate := "PIDData".D_ModeActivate, D_Mode := "PIDData".D_Mode, D_Interlock := "PIDData".D_Interlock, ChannelSelect := "PIDData".ChannelSelect, Setpoint => "ProcessData".PIDSetpoint, Input => "ProcessData".PIDInput, InputPER => "ProcessData".PIDInput_PER, ErrorACK => "ProcessData".PIDErrorAck, Reset => "ProcessData".PIDReset, ModeActivate => "ProcessData".PIDModeActivate, Mode => "ProcessData".PIDMode, Interlock => "ProcessData".PIDInterlock)
   END_RUNG
   // the same network as SCL:
   "PIDSwitch_DB"(A_Setpoint := "PIDData".A_Setpoint,   // "PIDSwitch"
                  A_Input := "PIDData".A_Input,
                  A_InputPER := "PIDData".A_InputPER,
                  A_ErrorACK := "PIDData".A_ErrorACK,
                  A_Reset := "PIDData".A_Reset,
                  A_ModeActivate := "PIDData".A_ModeActivate,
                  A_Mode := "PIDData".A_Mode,
                  A_Interlock := "PIDData".A_Interlock,
                  B_Setpoint := "PIDData".B_Setpoint,
                  B_Input := "PIDData".B_Input,
                  B_InputPER := "PIDData".B_InputPER,
                  B_ErrorACK := "PIDData".B_ErrorACK,
                  B_Reset := "PIDData".B_Reset,
                  B_ModeActivate := "PIDData".B_ModeActivate,
                  B_Mode := "PIDData".B_Mode,
                  B_Interlock := "PIDData".B_Interlock,
                  C_Setpoint := "PIDData".C_Setpoint,
                  C_Input := "PIDData".C_Input,
                  C_InputPER := "PIDData".C_InputPER,
                  C_ErrorACK := "PIDData".C_ErrorACK,
                  C_Reset := "PIDData".C_Reset,
                  C_ModeActivate := "PIDData".C_ModeActivate,
                  C_Mode := "PIDData".C_Mode,
                  C_Interlock := "PIDData".C_Interlock,
                  D_Setpoint := "PIDData".D_Setpoint,
                  D_Input := "PIDData".D_Input,
                  D_InputPER := "PIDData".A_InputPER,
                  D_ErrorACK := "PIDData".D_ErrorACK,
                  D_Reset := "PIDData".D_Reset,
                  D_ModeActivate := "PIDData".D_ModeActivate,
                  D_Mode := "PIDData".D_Mode,
                  D_Interlock := "PIDData".D_Interlock,
                  ChannelSelect := "PIDData".ChannelSelect,
                  Setpoint => "ProcessData".PIDSetpoint,
                  Input => "ProcessData".PIDInput,
                  InputPER => "ProcessData".PIDInput_PER,
                  ErrorACK => "ProcessData".PIDErrorAck,
                  Reset => "ProcessData".PIDReset,
                  ModeActivate => "ProcessData".PIDModeActivate,
                  Mode => "ProcessData".PIDMode,
                  Interlock => "ProcessData".PIDInterlock);
END_REGION

REGION Network 20: Beacon Light Green
   RUNG wire#powerrail
      Contact( "Operation".LampTest )
      Contact( "Clock_1Hz" )
      Coil( "BeaconLightGreen" )
   END_RUNG
   // the same network as SCL:
   "BeaconLightGreen" := "Operation".LampTest AND "Clock_1Hz";
END_REGION

REGION Network 21: Beacon Light Orange
   RUNG wire#powerrail
      Contact( "Operation".LampTest )
      wire#w1
      Contact( "Clock_1Hz" )
      Coil( "BeaconLightOrange" )
   END_RUNG
   RUNG wire#powerrail
      Contact( "Operation".RecruimentSignal )
   END_RUNG wire#w1
   RUNG wire#powerrail
      Contact( "Operation".RecruimentSignalEnding )
   END_RUNG wire#w1
   // the same network as SCL:
   "BeaconLightOrange" := ("Operation".LampTest OR "Operation".RecruimentSignal OR "Operation".RecruimentSignalEnding) AND "Clock_1Hz";
END_REGION

REGION Network 22: Beacon Light Red
   RUNG wire#powerrail
      Contact( "Operation".LampTest )
      Contact( "Clock_1Hz" )
      Coil( "BeaconLightRed" )
   END_RUNG
   // the same network as SCL:
   "BeaconLightRed" := "Operation".LampTest AND "Clock_1Hz";
END_REGION

